(* Logix 5000 project; controller PLC_MCC1300_75F1 vendor 1 type 14 code 166 rev 32.11; software revision 32.04; part 34 of 83 *)
(* tags used below, declared in another part *)
   C5 : COUNTER[51];
   CNV10_FLT : ALIAS FOR I[4].9;
   CNV10_FWD : ALIAS FOR O[5].9;
   CNV11_FLT : ALIAS FOR I[4].10;
   CNV11_FWD : ALIAS FOR O[5].10;
   CNV12_FLT : ALIAS FOR I[4].11;
   CNV1_FLT : ALIAS FOR I[4].0;
   CNV1_FWD : ALIAS FOR O[5].0;
   CNV2_FLT : ALIAS FOR I[4].1;
   CNV2_FWD : ALIAS FOR O[5].1;
   CNV3_FLT : ALIAS FOR I[4].2;
   CNV3_FWD : ALIAS FOR O[5].2;
   CNV4_FLT : ALIAS FOR I[4].3;
   CNV4_FWD : ALIAS FOR O[5].3;
   CNV5_FLT : ALIAS FOR I[4].4;
   CNV5_FWD : ALIAS FOR O[5].4;
   CNV6_FLT : ALIAS FOR I[4].5;
   CNV6_FWD : ALIAS FOR O[5].5;
   CNV7_FLT : ALIAS FOR I[4].6;
   CNV7_FWD : ALIAS FOR O[5].6;
   CNV8_FLT : ALIAS FOR I[4].7;
   CNV8_FWD : ALIAS FOR O[5].7;
   CNV9_FLT : ALIAS FOR I[4].8;
   CNV9_FWD : ALIAS FOR O[21].8;
   I : INT[128];   // Local Input Updates Input Slot 2
   N131 : INT[8];
   N14 : DINT[500];
   N803 : INT[420];
   O : INT[128];
   T4 : TIMER[51];
   T9 : TIMER[22];
(* MainProgram, continued *)

ROUTINE _75_LADDER   (* ladder *)
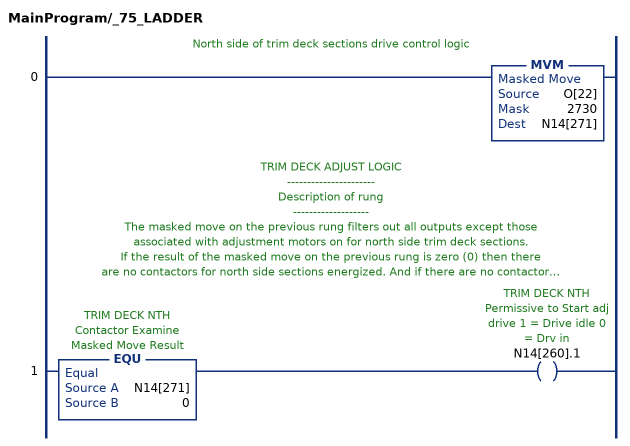
   // North side of trim deck sections drive control logic
   0: MVM(O[22],2730,N14[271]);
   // TRIM DECK ADJUST LOGIC
   // ----------------------
   // Description of rung
   // -------------------
   // The masked move on the previous rung filters out all outputs except those
   // associated with adjustment motors on for north side trim deck sections.
   // If the result of the masked move on the previous rung is zero (0) then there
   // are no contactors for north side sections energized. And if there are no contactors
   // for north side sections energized, then any north section may be energized.
   // As soon as the contactor for any section energizes, the result of the mased move on the
   // HISTORY
   // =======
   // DATE        DESCRIPTION                                                       PROGRAMMER
   // ====        ===========                                                       ==========
   // 2/29/96     Entered rung as designed                                          WAS
   // 3/1/96      Entered comment                                                   WAS
   1: EQU(N14[271],0)OTE(N14[260].1);
END_ROUTINE

ROUTINE _7_MCP_F   (* ladder *)
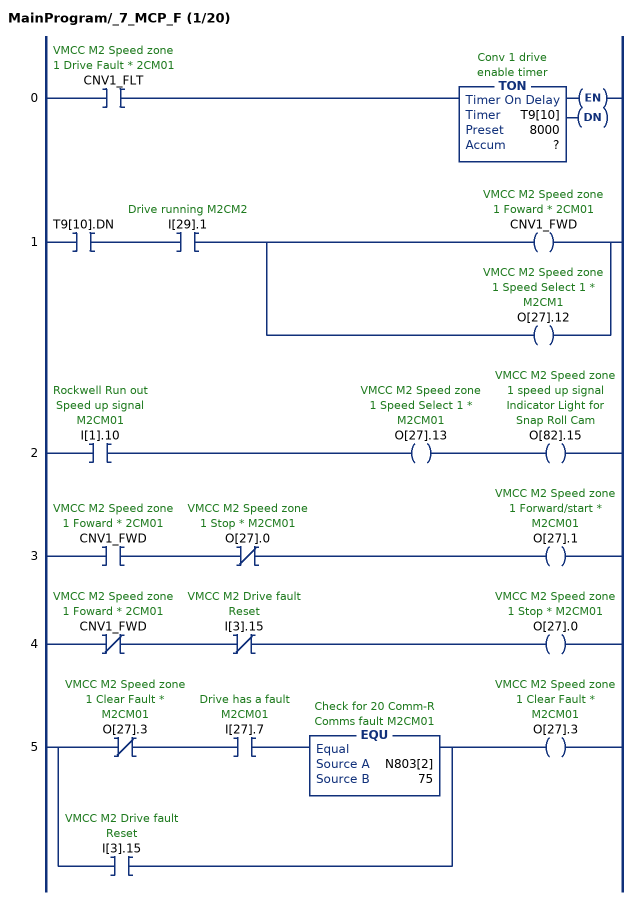
   0: XIC(CNV1_FLT)TON(T9[10],?,?);
   1: XIC(T9[10].DN)XIC(I[29].1)[OTE(CNV1_FWD) ,OTE(O[27].12) ];
   2: XIC(I[1].10)OTE(O[27].13)OTE(O[82].15);
   3: XIC(CNV1_FWD)XIO(O[27].0)OTE(O[27].1);
   4: XIO(CNV1_FWD)XIO(I[3].15)OTE(O[27].0);
   5: [XIO(O[27].3) XIC(I[27].7) EQU(N803[2],75) ,XIC(I[3].15) ]OTE(O[27].3);
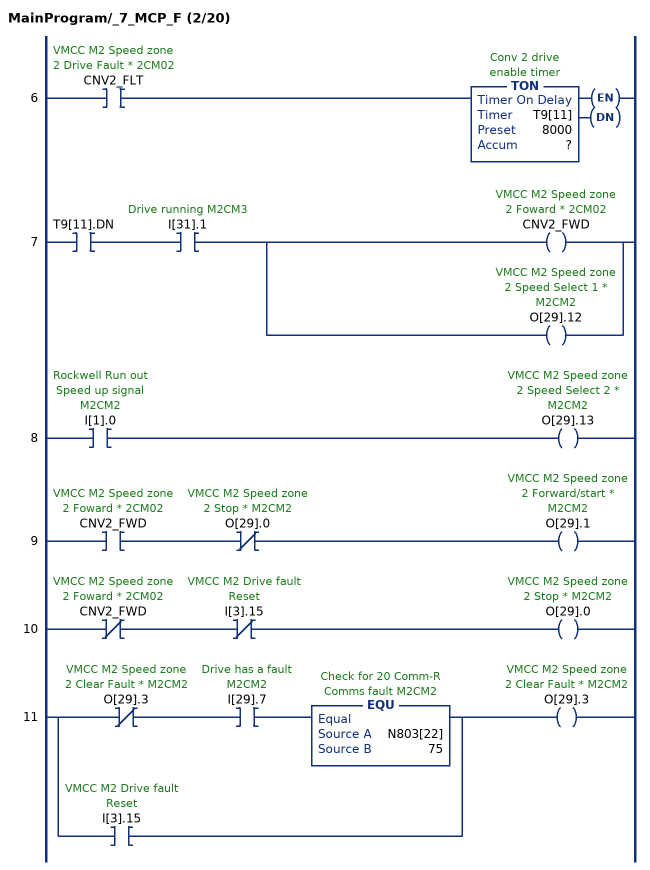
   6: XIC(CNV2_FLT)TON(T9[11],?,?);
   7: XIC(T9[11].DN)XIC(I[31].1)[OTE(CNV2_FWD) ,OTE(O[29].12) ];
   8: XIC(I[1].0)OTE(O[29].13);
   9: XIC(CNV2_FWD)XIO(O[29].0)OTE(O[29].1);
   10: XIO(CNV2_FWD)XIO(I[3].15)OTE(O[29].0);
   11: [XIO(O[29].3) XIC(I[29].7) EQU(N803[22],75) ,XIC(I[3].15) ]OTE(O[29].3);
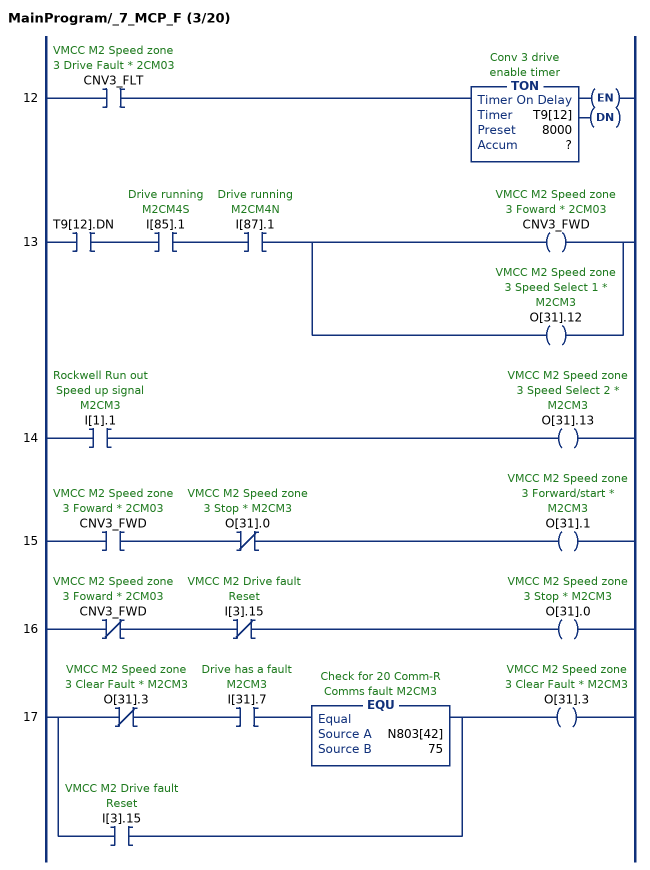
   12: XIC(CNV3_FLT)TON(T9[12],?,?);
   13: XIC(T9[12].DN)XIC(I[85].1)XIC(I[87].1)[OTE(CNV3_FWD) ,OTE(O[31].12) ];
   14: XIC(I[1].1)OTE(O[31].13);
   15: XIC(CNV3_FWD)XIO(O[31].0)OTE(O[31].1);
   16: XIO(CNV3_FWD)XIO(I[3].15)OTE(O[31].0);
   17: [XIO(O[31].3) XIC(I[31].7) EQU(N803[42],75) ,XIC(I[3].15) ]OTE(O[31].3);
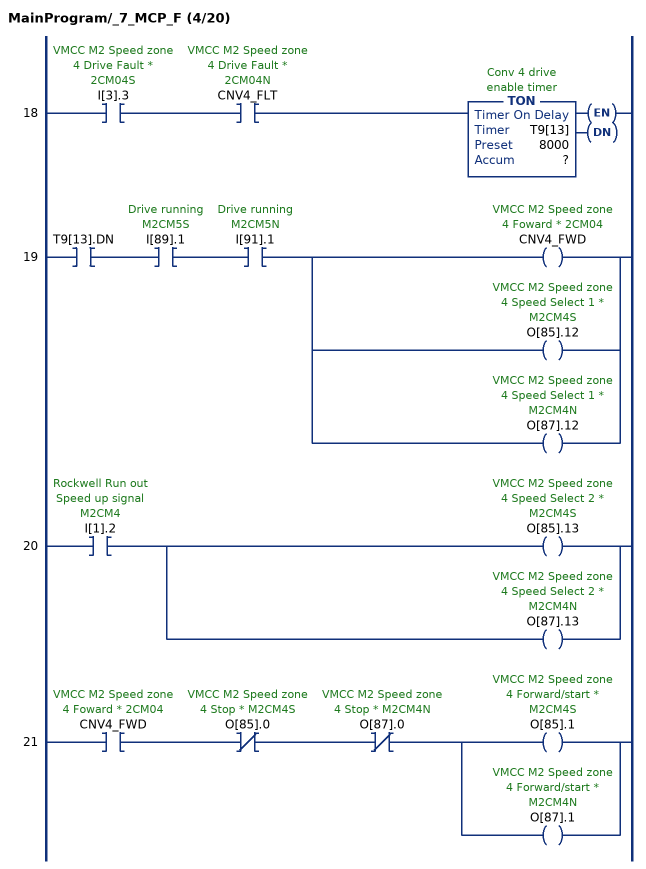
   18: XIC(I[3].3)XIC(CNV4_FLT)TON(T9[13],?,?);
   19: XIC(T9[13].DN)XIC(I[89].1)XIC(I[91].1)[OTE(CNV4_FWD) ,OTE(O[85].12) ,OTE(O[87].12) ];
   20: XIC(I[1].2)[OTE(O[85].13) ,OTE(O[87].13) ];
   21: XIC(CNV4_FWD)XIO(O[85].0)XIO(O[87].0)[OTE(O[85].1) ,OTE(O[87].1) ];
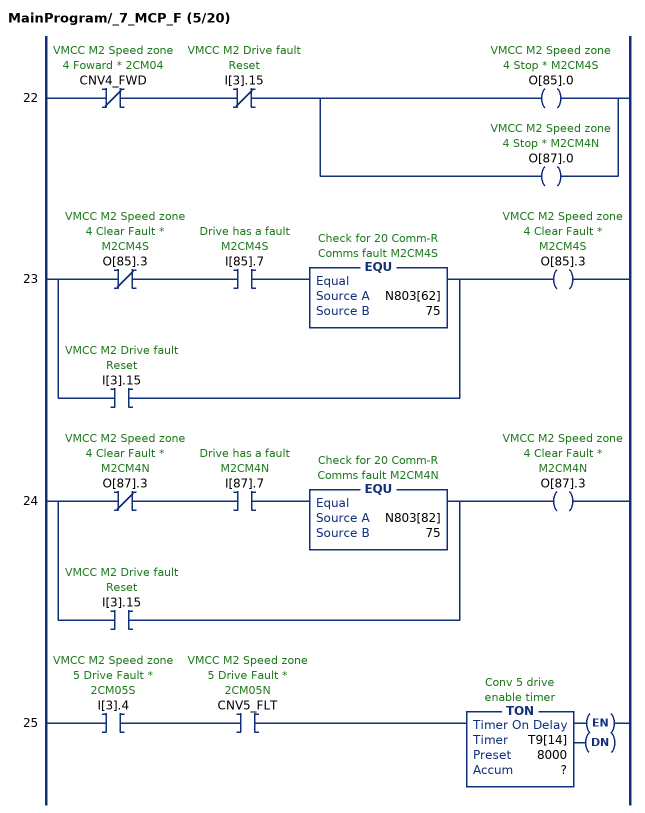
   22: XIO(CNV4_FWD)XIO(I[3].15)[OTE(O[85].0) ,OTE(O[87].0) ];
   23: [XIO(O[85].3) XIC(I[85].7) EQU(N803[62],75) ,XIC(I[3].15) ]OTE(O[85].3);
   24: [XIO(O[87].3) XIC(I[87].7) EQU(N803[82],75) ,XIC(I[3].15) ]OTE(O[87].3);
   25: XIC(I[3].4)XIC(CNV5_FLT)TON(T9[14],?,?);
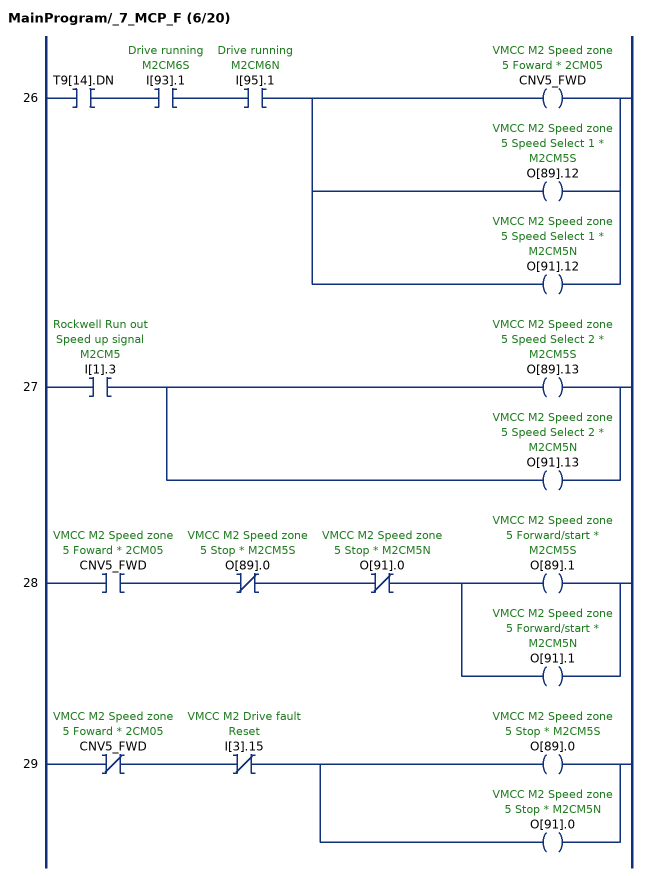
   26: XIC(T9[14].DN)XIC(I[93].1)XIC(I[95].1)[OTE(CNV5_FWD) ,OTE(O[89].12) ,OTE(O[91].12) ];
   27: XIC(I[1].3)[OTE(O[89].13) ,OTE(O[91].13) ];
   28: XIC(CNV5_FWD)XIO(O[89].0)XIO(O[91].0)[OTE(O[89].1) ,OTE(O[91].1) ];
   29: XIO(CNV5_FWD)XIO(I[3].15)[OTE(O[89].0) ,OTE(O[91].0) ];
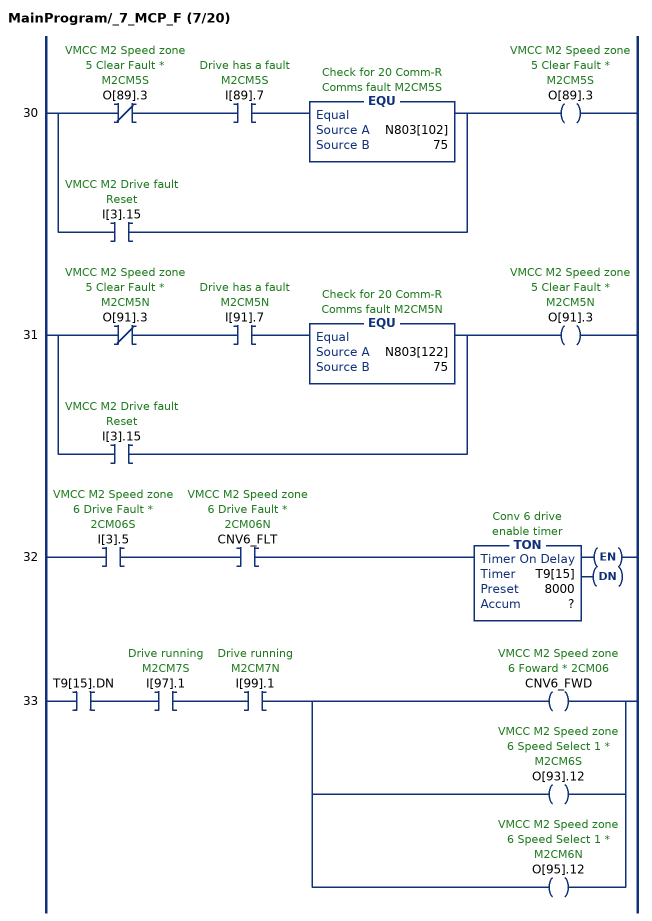
   30: [XIO(O[89].3) XIC(I[89].7) EQU(N803[102],75) ,XIC(I[3].15) ]OTE(O[89].3);
   31: [XIO(O[91].3) XIC(I[91].7) EQU(N803[122],75) ,XIC(I[3].15) ]OTE(O[91].3);
   32: XIC(I[3].5)XIC(CNV6_FLT)TON(T9[15],?,?);
   33: XIC(T9[15].DN)XIC(I[97].1)XIC(I[99].1)[OTE(CNV6_FWD) ,OTE(O[93].12) ,OTE(O[95].12) ];
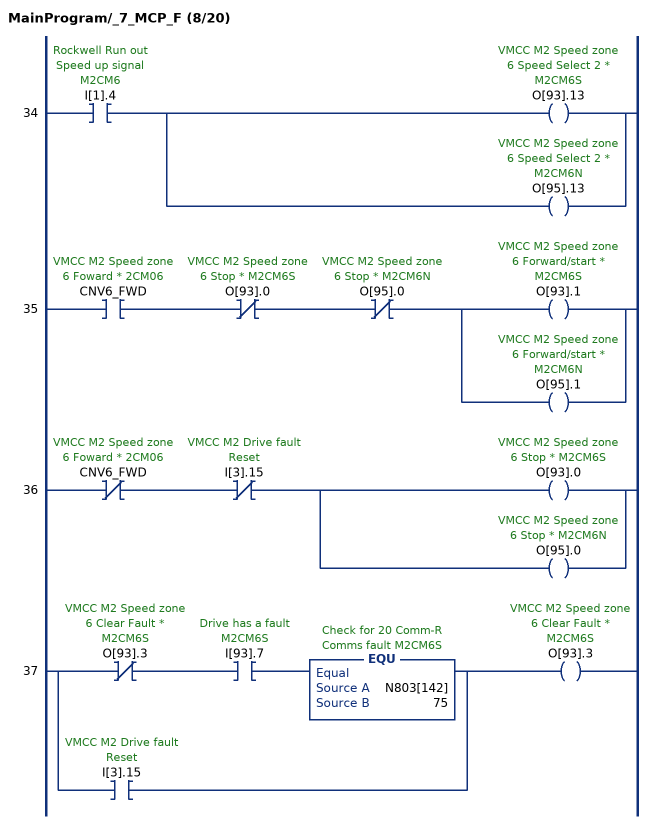
   34: XIC(I[1].4)[OTE(O[93].13) ,OTE(O[95].13) ];
   35: XIC(CNV6_FWD)XIO(O[93].0)XIO(O[95].0)[OTE(O[93].1) ,OTE(O[95].1) ];
   36: XIO(CNV6_FWD)XIO(I[3].15)[OTE(O[93].0) ,OTE(O[95].0) ];
   37: [XIO(O[93].3) XIC(I[93].7) EQU(N803[142],75) ,XIC(I[3].15) ]OTE(O[93].3);
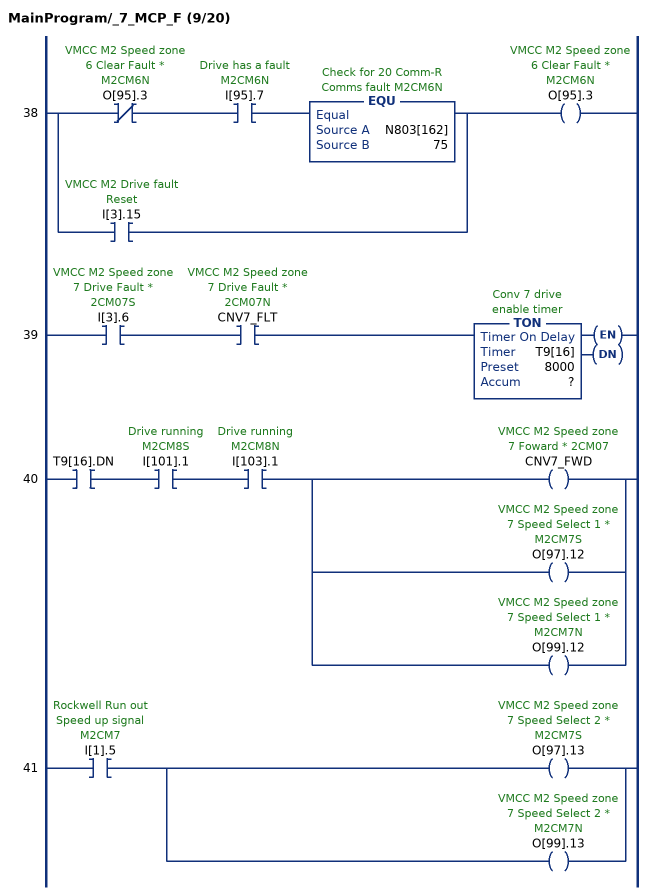
   38: [XIO(O[95].3) XIC(I[95].7) EQU(N803[162],75) ,XIC(I[3].15) ]OTE(O[95].3);
   39: XIC(I[3].6)XIC(CNV7_FLT)TON(T9[16],?,?);
   40: XIC(T9[16].DN)XIC(I[101].1)XIC(I[103].1)[OTE(CNV7_FWD) ,OTE(O[97].12) ,OTE(O[99].12) ];
   41: XIC(I[1].5)[OTE(O[97].13) ,OTE(O[99].13) ];
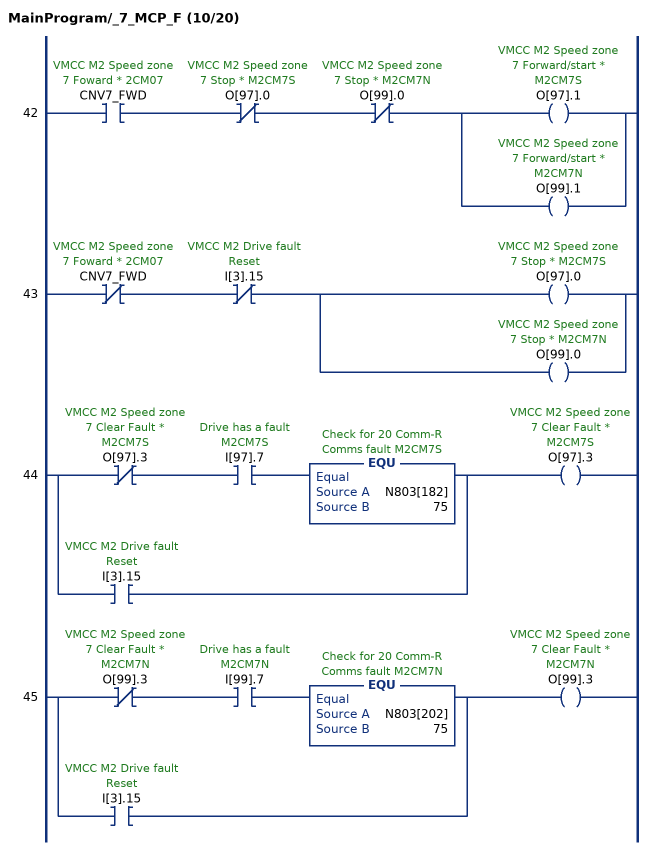
   42: XIC(CNV7_FWD)XIO(O[97].0)XIO(O[99].0)[OTE(O[97].1) ,OTE(O[99].1) ];
   43: XIO(CNV7_FWD)XIO(I[3].15)[OTE(O[97].0) ,OTE(O[99].0) ];
   44: [XIO(O[97].3) XIC(I[97].7) EQU(N803[182],75) ,XIC(I[3].15) ]OTE(O[97].3);
   45: [XIO(O[99].3) XIC(I[99].7) EQU(N803[202],75) ,XIC(I[3].15) ]OTE(O[99].3);
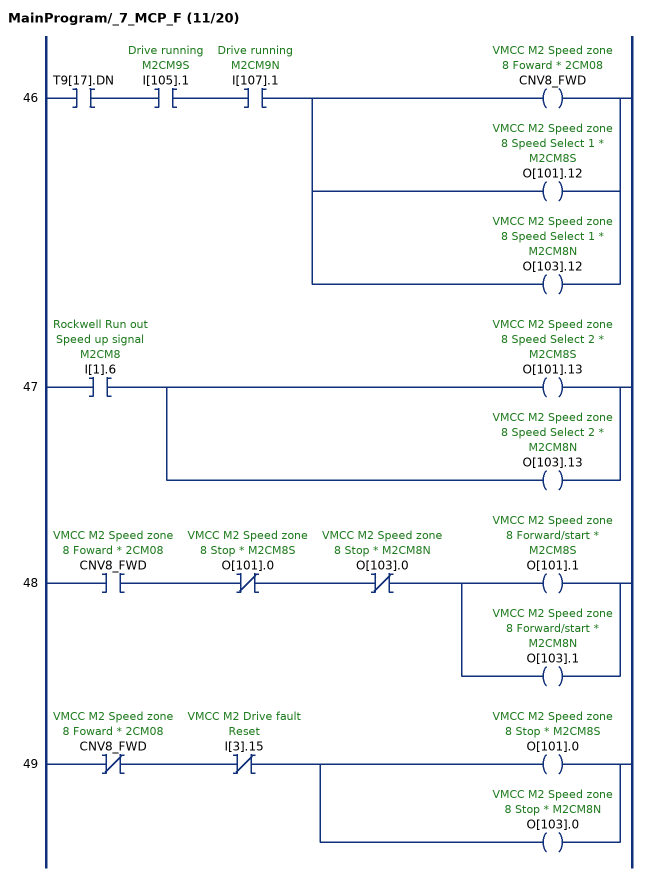
   46: XIC(T9[17].DN)XIC(I[105].1)XIC(I[107].1)[OTE(CNV8_FWD) ,OTE(O[101].12) ,OTE(O[103].12) ];
   47: XIC(I[1].6)[OTE(O[101].13) ,OTE(O[103].13) ];
   48: XIC(CNV8_FWD)XIO(O[101].0)XIO(O[103].0)[OTE(O[101].1) ,OTE(O[103].1) ];
   49: XIO(CNV8_FWD)XIO(I[3].15)[OTE(O[101].0) ,OTE(O[103].0) ];
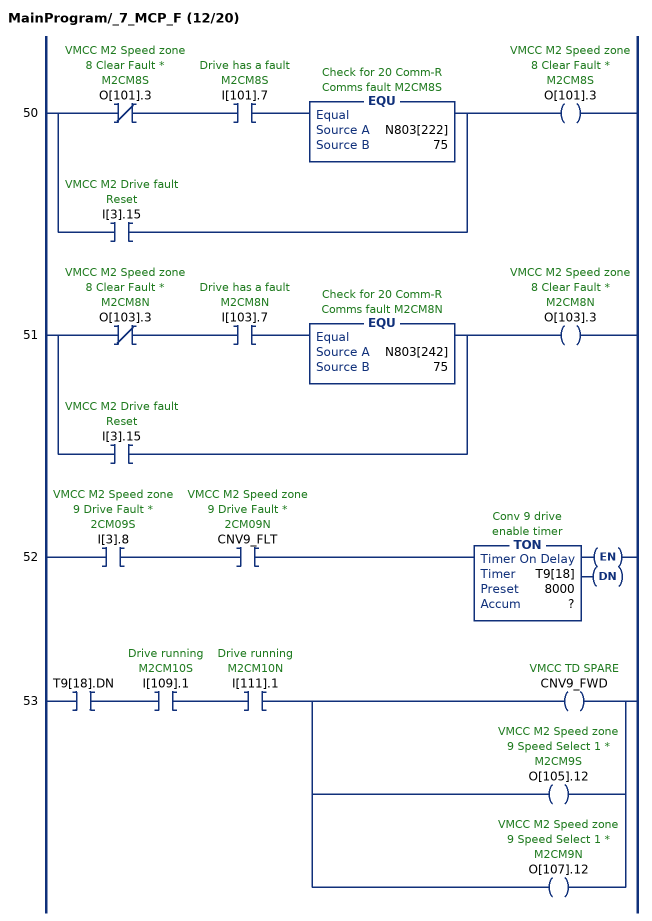
   50: [XIO(O[101].3) XIC(I[101].7) EQU(N803[222],75) ,XIC(I[3].15) ]OTE(O[101].3);
   51: [XIO(O[103].3) XIC(I[103].7) EQU(N803[242],75) ,XIC(I[3].15) ]OTE(O[103].3);
   52: XIC(I[3].8)XIC(CNV9_FLT)TON(T9[18],?,?);
   53: XIC(T9[18].DN)XIC(I[109].1)XIC(I[111].1)[OTE(CNV9_FWD) ,OTE(O[105].12) ,OTE(O[107].12) ];
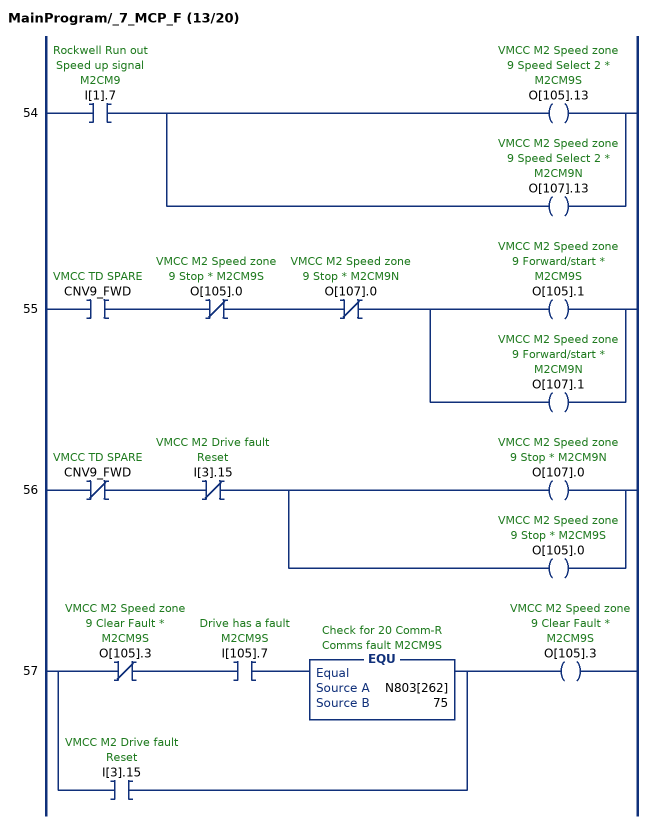
   54: XIC(I[1].7)[OTE(O[105].13) ,OTE(O[107].13) ];
   55: XIC(CNV9_FWD)XIO(O[105].0)XIO(O[107].0)[OTE(O[105].1) ,OTE(O[107].1) ];
   56: XIO(CNV9_FWD)XIO(I[3].15)[OTE(O[107].0) ,OTE(O[105].0) ];
   57: [XIO(O[105].3) XIC(I[105].7) EQU(N803[262],75) ,XIC(I[3].15) ]OTE(O[105].3);
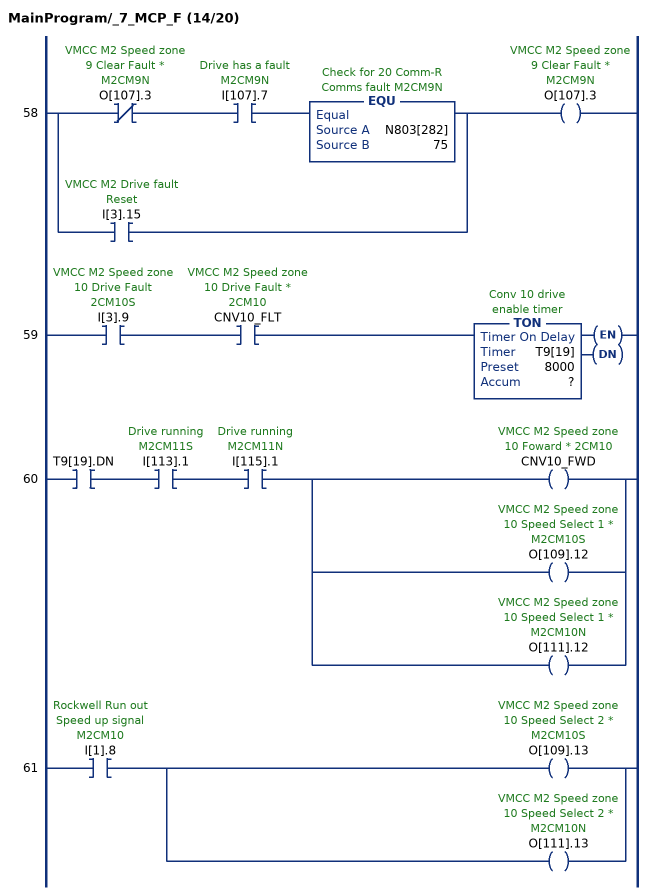
   58: [XIO(O[107].3) XIC(I[107].7) EQU(N803[282],75) ,XIC(I[3].15) ]OTE(O[107].3);
   59: XIC(I[3].9)XIC(CNV10_FLT)TON(T9[19],?,?);
   60: XIC(T9[19].DN)XIC(I[113].1)XIC(I[115].1)[OTE(CNV10_FWD) ,OTE(O[109].12) ,OTE(O[111].12) ];
   61: XIC(I[1].8)[OTE(O[109].13) ,OTE(O[111].13) ];
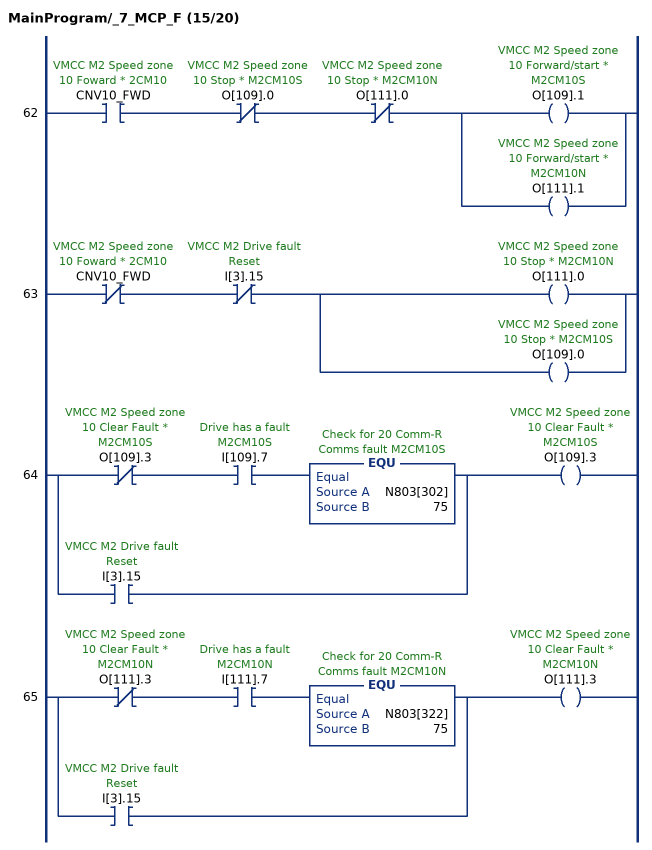
   62: XIC(CNV10_FWD)XIO(O[109].0)XIO(O[111].0)[OTE(O[109].1) ,OTE(O[111].1) ];
   63: XIO(CNV10_FWD)XIO(I[3].15)[OTE(O[111].0) ,OTE(O[109].0) ];
   64: [XIO(O[109].3) XIC(I[109].7) EQU(N803[302],75) ,XIC(I[3].15) ]OTE(O[109].3);
   65: [XIO(O[111].3) XIC(I[111].7) EQU(N803[322],75) ,XIC(I[3].15) ]OTE(O[111].3);
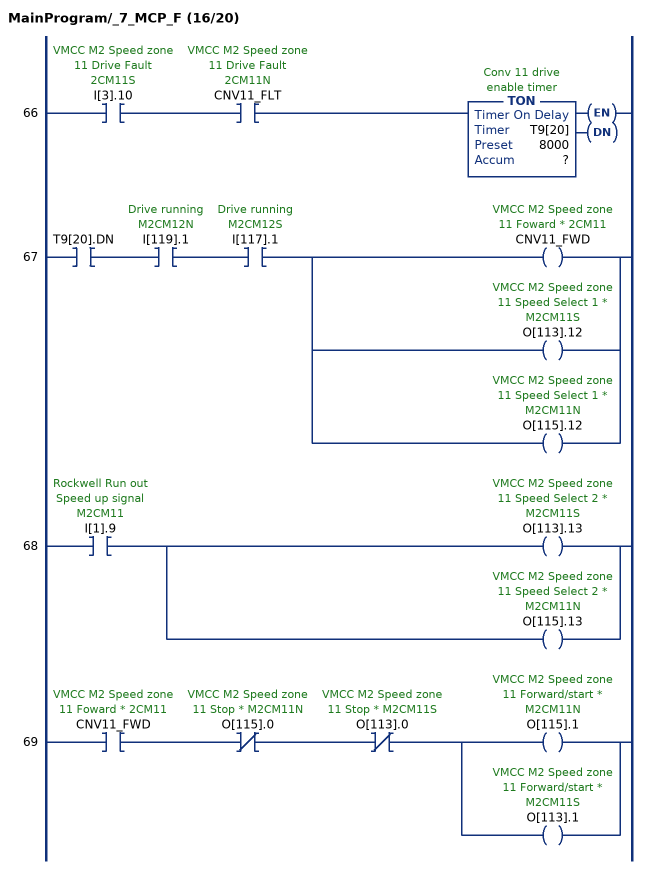
   66: XIC(I[3].10)XIC(CNV11_FLT)TON(T9[20],?,?);
   67: XIC(T9[20].DN)XIC(I[119].1)XIC(I[117].1)[OTE(CNV11_FWD) ,OTE(O[113].12) ,OTE(O[115].12) ];
   68: XIC(I[1].9)[OTE(O[113].13) ,OTE(O[115].13) ];
   69: XIC(CNV11_FWD)XIO(O[115].0)XIO(O[113].0)[OTE(O[115].1) ,OTE(O[113].1) ];
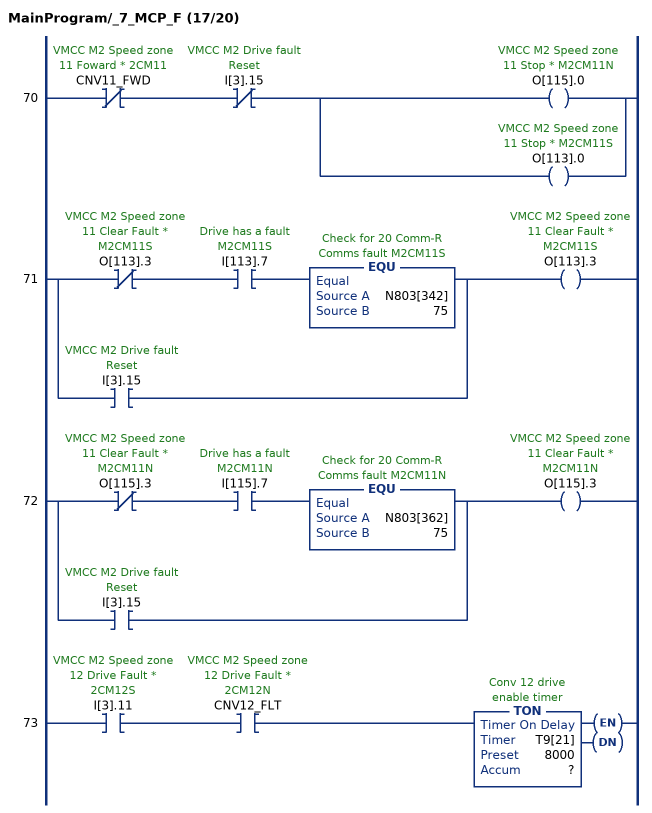
   70: XIO(CNV11_FWD)XIO(I[3].15)[OTE(O[115].0) ,OTE(O[113].0) ];
   71: [XIO(O[113].3) XIC(I[113].7) EQU(N803[342],75) ,XIC(I[3].15) ]OTE(O[113].3);
   72: [XIO(O[115].3) XIC(I[115].7) EQU(N803[362],75) ,XIC(I[3].15) ]OTE(O[115].3);
   73: XIC(I[3].11)XIC(CNV12_FLT)TON(T9[21],?,?);
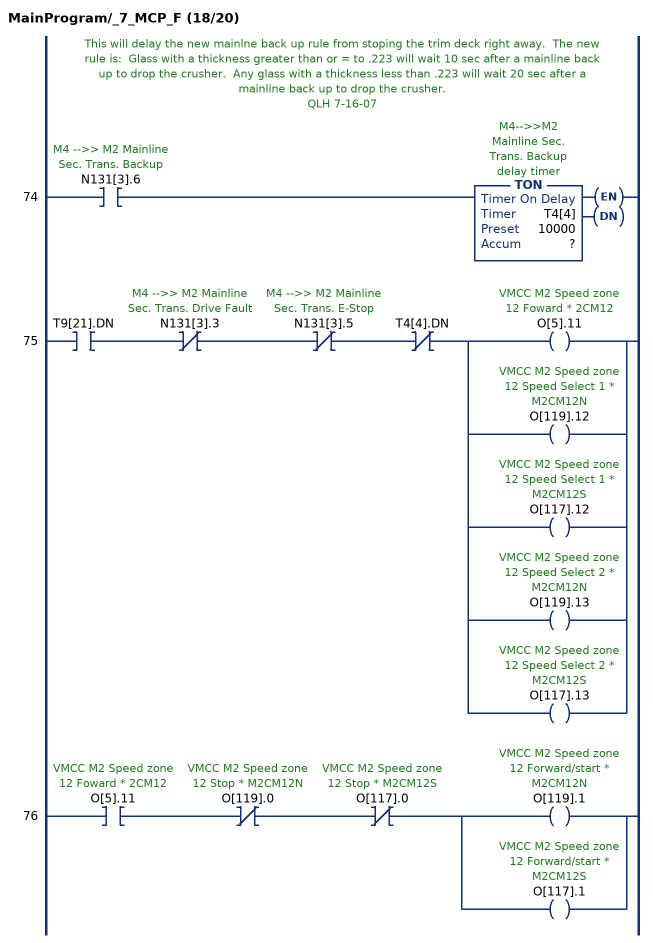
   // This will delay the new mainlne back up rule from stoping the trim deck right away.  The new rule is:  Glass with a thickness greater than or = to .223 will wait 10 sec after a mainline back up to drop the crusher.  Any glass with a thickness less than .223 will wait 20 sec after a mainline back up to drop the crusher.
   // QLH 7-16-07
   74: XIC(N131[3].6)TON(T4[4],?,?);
   75: XIC(T9[21].DN)XIO(N131[3].3)XIO(N131[3].5)XIO(T4[4].DN)[OTE(O[5].11) ,OTE(O[119].12) ,OTE(O[117].12) ,OTE(O[119].13) ,OTE(O[117].13) ];
   76: XIC(O[5].11)XIO(O[119].0)XIO(O[117].0)[OTE(O[119].1) ,OTE(O[117].1) ];
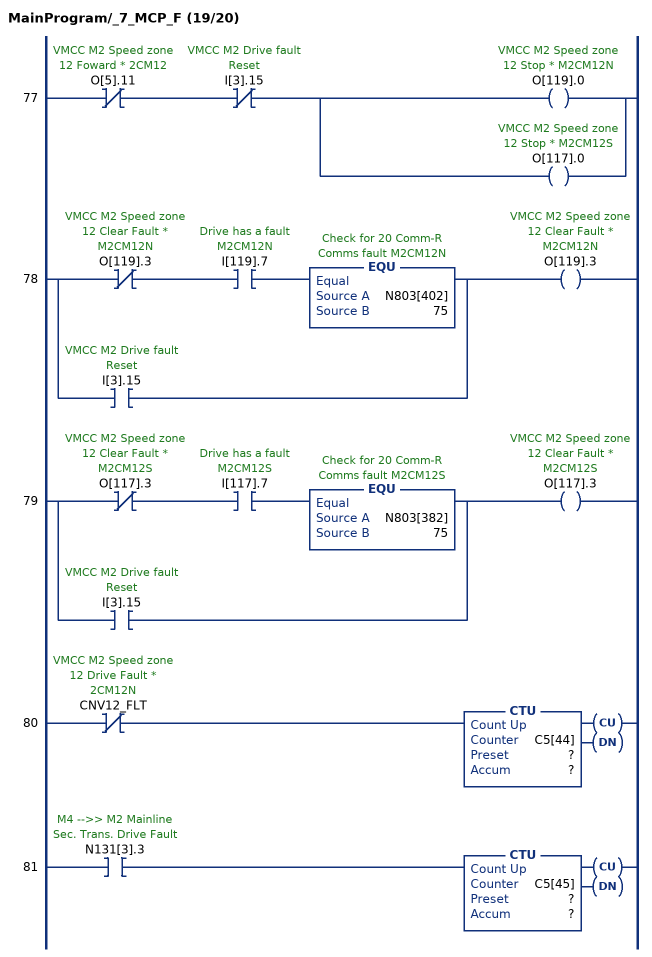
   77: XIO(O[5].11)XIO(I[3].15)[OTE(O[119].0) ,OTE(O[117].0) ];
   78: [XIO(O[119].3) XIC(I[119].7) EQU(N803[402],75) ,XIC(I[3].15) ]OTE(O[119].3);
   79: [XIO(O[117].3) XIC(I[117].7) EQU(N803[382],75) ,XIC(I[3].15) ]OTE(O[117].3);
   80: XIO(CNV12_FLT)CTU(C5[44],?,?);
   81: XIC(N131[3].3)CTU(C5[45],?,?);
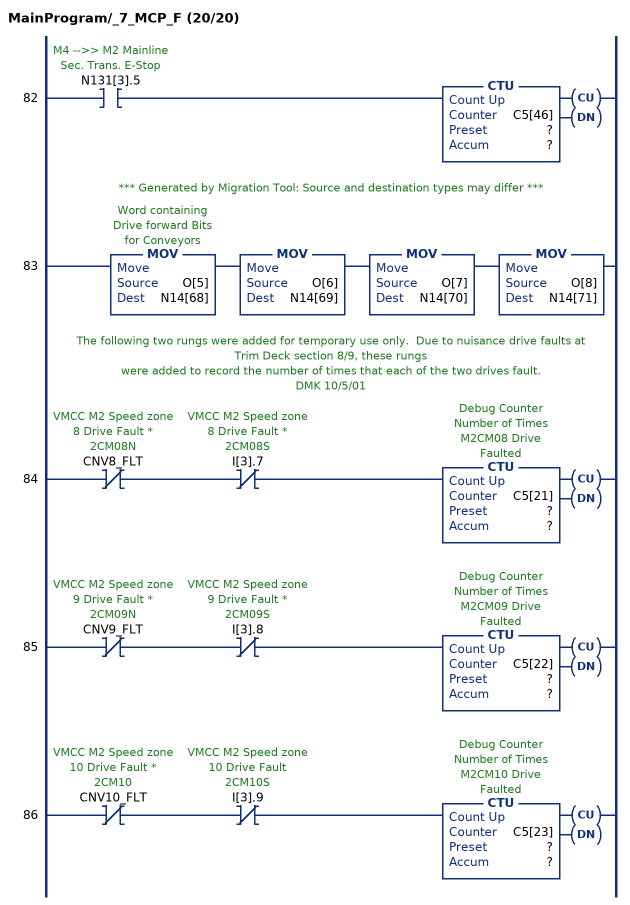
   82: XIC(N131[3].5)CTU(C5[46],?,?);
   // *** Generated by Migration Tool: Source and destination types may differ ***
   83: MOV(O[5],N14[68])MOV(O[6],N14[69])MOV(O[7],N14[70])MOV(O[8],N14[71]);
   // The following two rungs were added for temporary use only.  Due to nuisance drive faults at Trim Deck section 8/9, these rungs
   // were added to record the number of times that each of the two drives fault.
   // DMK 10/5/01
   84: XIO(CNV8_FLT)XIO(I[3].7)CTU(C5[21],?,?);
   85: XIO(CNV9_FLT)XIO(I[3].8)CTU(C5[22],?,?);
   86: XIO(CNV10_FLT)XIO(I[3].9)CTU(C5[23],?,?);
END_ROUTINE
